(* Logix 5000 project; controller PLC_MCC1300_75F1 vendor 1 type 14 code 166 rev 32.11; software revision 32.04; part 4 of 83 *)
(* tags used below, declared in another part *)
   GP_AccTimeForGap : GP_AccTimeForGap;
   GP_CheckIdPlatePresent : GP_CheckIdPlatePresent;
   GP_ConversionXY : GP_ConversionXY;
   GP_ConvertDataFromStacker : GP_ConvertDataFromStacker;
   GP_ConvertDataToStacker : GP_ConvertDataToStacker;
   GP_InvertCapxLite : GP_InvertCapxLite;

ADD_ON_INSTRUCTION GP_AccTimeForGap   (* revision 1.0 *)
VAR_INPUT
   IN_dLehrSpeed_mm_min : DINT; {access None, required}
   IN_dLineSpeed_mm_min : DINT; {access None, required}
   IN_rAcc_m_s2 : REAL; {access None, required}
   IN_dGapRequested_cmm : DINT; {access None, required}
END_VAR
VAR_OUTPUT
   OUT_dAccTime_ms : DINT; {access None, required}
END_VAR
VAR
   TMP_rSpeed_mm_s : REAL; {access None}
   TMP_rConvSpeed_mm_s : REAL; {access None}
   TMP_rAccConv_mm_s2 : REAL; {access None}
   TMP_rAcc : REAL; {access None}
   TMP_rSv : REAL; {access None}
   TMP_dGap_mm : DINT; {access None}
END_VAR

ROUTINE Logic   (* structured text *)
   
   TMP_rSpeed_mm_s := (IN_dLehrSpeed_mm_min / 60.0);
   TMP_rConvSpeed_mm_s := (IN_dLineSpeed_mm_min / 60.0);
   TMP_rAccConv_mm_s2 := (IN_rAcc_m_s2 * 1000.0);
   TMP_dGap_mm := (IN_dGapRequested_cmm / 100);
   
   TMP_rAcc := ((TMP_rSpeed_mm_s*-1) + SQRT(TMP_rSpeed_mm_s**2 + (2*TMP_rAccConv_mm_s2*200)))/TMP_rAccConv_mm_s2;
   IF ((TMP_rAcc*TMP_rAccConv_mm_s2) + TMP_rSpeed_mm_s) > TMP_rConvSpeed_mm_s THEN
       TMP_rAcc := (TMP_rConvSpeed_mm_s - TMP_rSpeed_mm_s) / TMP_rAccConv_mm_s2;
       TMP_rSv := TMP_dGap_mm - (0.5*(TMP_rAcc**2)*TMP_rAccConv_mm_s2) - (TMP_rSpeed_mm_s*TMP_rAcc);
       TMP_rAcc := TMP_rAcc + (TMP_rSv/TMP_rConvSpeed_mm_s);
   END_IF;
   
   IF IN_dGapRequested_cmm > 0 THEN
       OUT_dAccTime_ms := TMP_rAcc * 1000.0;
   ELSE
       OUT_dAccTime_ms := 0;
   END_IF;
   
END_ROUTINE
END_ADD_ON_INSTRUCTION

ADD_ON_INSTRUCTION GP_BaricenterDefinition   (* revision 1.0 *)
VAR_INPUT
   In_dHeadPosition : DINT; {required}   // Head position on conveyor below [mm/100]
END_VAR
VAR_IN_OUT
   InOut_ConvoyData : UDT_Convoy_SL; {required}
END_VAR
VAR_INPUT
   In_dInLitePos : DINT; {access None, required}   // Position input lite - Left to Right line flow(0=AX; 1=XA)
   In_dOutDirection : DINT; {required}   // Direction of lateral flow (0=Left; 1=Right; 2=CW(rotation); 3=CCW(rotation))
   In_dOutLitePos : DINT; {access None, required}   // Position output lite - Left to Right line flow(0=AX; 1=XA)
   In_dOffset1 : DINT; {required}   // Distance of start conveyorIn and axe conveyorOut [mm/100]
   In_dOffset2 : DINT; {required}   // (NU)
   In_dConveyorLenght : DINT; {access None, required}   // Conveyor below [mm/100]
   In_dConveyorWidth : DINT; {access None, required}   // Conveyor below [mm/100]
END_VAR
VAR
   TMP_idxCap : DINT; {access None}
   TMP_IdxLite : DINT; {access None}
   TMP_MaxCap : DINT; {access None}
   TMP_MaxLite : DINT; {access None}
   TMP_d : DINT; {access None}
   TMP_NewBarycenterCap : DINT[10]; {access None}
   TMP_HeadPosition : DINT[10]; {access None}   // Head position cap [mm/100]
END_VAR

ROUTINE Logic   (* structured text *)
   ////////////////////////////////////////////////////////////
   //   Copyright (c)  <Key Automation srl>
   //------------------------------------------------------------
   //   Routine: GP_BaricenterDefinition - Logic
   //   Author: Gerto\admin
   //   Created: 2020-02-06
   //------------------------------------------------------------
   //   Description:
   //
   //
   //   History:
   //
   ////////////////////////////////////////////////////////////
   
   //Dimension array
   Size(InOut_ConvoyData.rgtCap,0,TMP_MaxCap);
   size(InOut_ConvoyData.rgtCap[0].rgtLite,0,TMP_MaxLite);
   
   //Conveyor deviation *****************************************
   
   //Cap1 Barycenter = HeadPosIn - 1/2 cap1lenght - offset1(distance between start of conveyorIn and exe of conveyorOut)
   //Cap2 Barycenter = Cap1 Barycenter - 1/2 Cap1Lenght - Gap - 1/2 Cap2Lenght
   //Cap3...
   if 	(In_dOutDirection = 0 and In_dInLitePos = 0 and In_dOutLitePos = 0) or
   	(In_dOutDirection = 0 and In_dInLitePos = 1 and In_dOutLitePos = 0) or
   	(In_dOutDirection = 1 and In_dInLitePos = 0 and In_dOutLitePos = 1) or
   	(In_dOutDirection = 1 and In_dInLitePos = 1 and In_dOutLitePos = 1) then
   	//Barycenter 1° cap
   	TMP_NewBarycenterCap[0] := In_dHeadPosition - InOut_ConvoyData.rgtCap[0].dLength_cmm/2 - In_dOffset1;
   	//Baricenter other caps
   	for TMP_idxCap := 1 to InOut_ConvoyData.dTotalCaps - 1 by 1 do
   		TMP_NewBarycenterCap[TMP_idxCap] := TMP_NewBarycenterCap[TMP_idxCap-1] - InOut_ConvoyData.rgtCap[TMP_idxCap-1].dLength_cmm / 2 - InOut_ConvoyData.rgtCap[TMP_idxCap-1].dReqGapForConv_cmm - InOut_ConvoyData.rgtCap[TMP_idxCap].dLength_cmm / 2;
   	end_for;
   end_if;
   
   
   //Cap1 Barycenter = - (head pos In - 1/2 Cap1Lenght - Offset1)
   //Cap2 Barycenter = Cap1 Barycenter + 1/2 Cap1Lenght + Gap + 1/2 Cap2Lenght-
   //Cap3...
   if 	(In_dOutDirection = 0 and In_dInLitePos = 0 and In_dOutLitePos = 1) or
   	(In_dOutDirection = 0 and In_dInLitePos = 1 and In_dOutLitePos = 1) or
   	(In_dOutDirection = 1 and In_dInLitePos = 0 and In_dOutLitePos = 0) or
   	(In_dOutDirection = 1 and In_dInLitePos = 1 and In_dOutLitePos = 0) then
   	//Baricenter 1° cap
   	TMP_NewBarycenterCap[0] := - (In_dHeadPosition - InOut_ConvoyData.rgtCap[0].dLength_cmm / 2 - In_dOffset1);
   	//Barycenter other caps
   	for TMP_idxCap := 1 to InOut_ConvoyData.dTotalCaps - 1 by 1 do
   		TMP_NewBarycenterCap[TMP_idxCap] := TMP_NewBarycenterCap[TMP_idxCap-1] + InOut_ConvoyData.rgtCap[TMP_idxCap-1].dLength_cmm / 2 + InOut_ConvoyData.rgtCap[TMP_idxCap-1].dReqGapForConv_cmm + InOut_ConvoyData.rgtCap[TMP_idxCap].dLength_cmm / 2;
   	end_for;
   end_if;
   
   
   //Rotator ****************************************************
   
   //Definition head position for all caps
   TMP_HeadPosition[0] := In_dHeadPosition;
   for TMP_idxCap := 1 to InOut_ConvoyData.dTotalCaps - 1 by 1 do
   	TMP_HeadPosition[TMP_idxCap] := TMP_HeadPosition[TMP_idxCap-1] - InOut_ConvoyData.rgtCap[TMP_idxCap-1].dLength_cmm - InOut_ConvoyData.rgtCap[TMP_idxCap-1].dReqGapForConv_cmm;
   end_for;
   
   
   //Cap[cap] Barycenter = (HeadPosCap[cap] - ConveyorLengthIn/2 - CapLength[cap]/2)
   if 	(In_dOutDirection = 2 and In_dInLitePos = 0 and In_dOutLitePos = 0) or
   	(In_dOutDirection = 3 and In_dInLitePos = 1 and In_dOutLitePos = 1) then
   	for TMP_idxCap := 0 to InOut_ConvoyData.dTotalCaps - 1 by 1 do
   		TMP_NewBarycenterCap[TMP_idxCap] := (TMP_HeadPosition[TMP_idxCap] - In_dConveyorLenght/2 - InOut_ConvoyData.rgtCap[TMP_idxCap].dLength_cmm/2);
   	end_for;
   end_if;
   
   //Cap[cap] Barycenter = - (HeadPosCap[cap] - ConveyorLengthIn/2 - CapLength[cap]/2)
   if 	(In_dOutDirection = 2 and In_dInLitePos = 1 and In_dOutLitePos = 1) or
   	(In_dOutDirection = 3 and In_dInLitePos = 0 and In_dOutLitePos = 0) then
   	for TMP_idxCap := 0 to InOut_ConvoyData.dTotalCaps - 1 by 1 do
   		TMP_NewBarycenterCap[TMP_idxCap] := -(TMP_HeadPosition[TMP_idxCap] - In_dConveyorLenght/2 - InOut_ConvoyData.rgtCap[TMP_idxCap].dLength_cmm/2);
   	end_for;
   end_if;
   
   //Write output
   for TMP_idxCap := 0 to InOut_ConvoyData.dTotalCaps - 1 by 1 do
   	for TMP_IdxLite := 0 to TMP_MaxLite - 1 by 1 do
   		if InOut_ConvoyData.rgtCap[TMP_idxCap].rgtLite[TMP_IdxLite].dID <> 0 then
   			InOut_ConvoyData.rgtCap[TMP_idxCap].rgtLite[TMP_IdxLite].dBarycenter_cmm := TMP_NewBarycenterCap[TMP_idxCap];
   		end_if;
   	end_for;
   end_for;
END_ROUTINE
END_ADD_ON_INSTRUCTION

ADD_ON_INSTRUCTION GP_CalculatePlateNumber   (* revision 1.0 *)
VAR_IN_OUT
   INO_tPlate : UDT_ConvoyCap_ZC; {required}   // Plate data
END_VAR
VAR
   TMP_dLiteSize : DINT; {access None}
   TMP_dLite : DINT; {access None}
   TMP_dCapSize : DINT; {access None}
   TMP_dCap : DINT; {access None}
   TMP_dCountCaps : DINT; {access None}
   TMP_dCountLites : DINT; {access None}
END_VAR

ROUTINE Logic   (* structured text *)
   //Initialize
   size(INO_tPlate.rgtCap[0],0,TMP_dCapSize);
   size(INO_tPlate.rgtCap[0].rgtLite[0],0,TMP_dLiteSize);
   
   TMP_dCountCaps:= 0;
   
   FOR TMP_dCap:= 0 TO TMP_dCapSize - 1 DO
   	TMP_dCountLites:= 0;
   	FOR TMP_dLite := 0 TO TMP_dLiteSize - 1 DO
   
   		IF INO_tPlate.rgtCap[TMP_dCap].rgtLite[TMP_dLite].dID <> 0 THEN
   
   			TMP_dCountLites := TMP_dCountLites +1 ;
   
   		END_IF;
   
   	END_FOR;
   
   	INO_tPlate.rgtCap[TMP_dCap].dNumLites := TMP_dCountLites ;
   
   	IF TMP_dCountLites > 0 THEN
   
   		TMP_dCountCaps := TMP_dCountCaps + 1 ;
   
   	END_IF;
   
   END_FOR;
   
   IF TMP_dCountCaps > 1 THEN
   
   	INO_tPlate.dTotalCaps := TMP_dCountCaps ;
   
   ELSE
   
   	INO_tPlate.dTotalCaps := 0 ;
   
   END_IF;
   
   EnableOut := 1 ;
END_ROUTINE
END_ADD_ON_INSTRUCTION

ADD_ON_INSTRUCTION GP_CheckIdAndDestination   (* revision 1.0 *)
VAR_INPUT
   IN_dDestMask1 : DINT; {access None, required}   // Destinations available on operator side
   IN_dDestMask2 : DINT; {access None, required}   // Destinations available on opposite operator side
END_VAR
VAR_IN_OUT
   INO_tPlate : UDT_Convoy_SL; {required}   // Plate data
   INO_rgxId : DINT[4]; {required}   // Array Id Plate present [Cap, Lite]
END_VAR
VAR_OUTPUT
   OUT_xIDPresent : BOOL; {access None}   // Id present
   OUT_xDest1Found : BOOL; {access None}   // Destinations found
   OUT_xDest2Found : BOOL; {access None}   // Destinations found
   OUT_xAlternative1Found : BOOL; {access None}   // Alternatives found
   OUT_xAlternative2Found : BOOL; {access None}   // Alternatives found
   OUT_x2Choice1Found : BOOL; {access None}   // 2°Choice found
   OUT_x2Choice2Found : BOOL; {access None}   // 2°Choice found
END_VAR
VAR
   TMP_dCap : DINT; {access None}
   TMP_dLite : DINT; {access None}
   TMP_dLiteSize : DINT; {access None}
   TMP_dCapSize : DINT; {access None}
END_VAR

ROUTINE Logic   (* structured text *)
   //Initialize
   INO_rgxId[0]:= 0; INO_rgxId[1]:= 0; INO_rgxId[2]:= 0;INO_rgxId[3]:= 0;
   OUT_xIDPresent:= 0;
   OUT_xDest1Found:= 0;
   OUT_xDest2Found:= 0;
   OUT_xAlternative1Found:= 0;
   OUT_xAlternative2Found:= 0;
   OUT_x2Choice1Found:= 0;
   OUT_x2Choice2Found:= 0;
   
   size(INO_tPlate.rgtCap[0],0,TMP_dCapSize);
   size(INO_tPlate.rgtCap[0].rgtLite[0],0,TMP_dLiteSize);
   
   //This function check ID Plate present
   //Max Cap = 4
   //Max Lite = 8
   FOR TMP_dCap:= 0 TO TMP_dCapSize - 1 DO
   
   	FOR TMP_dLite := 0 TO TMP_dLiteSize - 1 DO
   
   	IF INO_tPlate.rgtCap[TMP_dCap].rgtLite[TMP_dLite].dID <> 0 THEN
   
   		OUT_xIDPresent:= 1;
   		INO_rgxId[TMP_dCap].[TMP_dLite]:= 1;
   		//Find available destination
   		IF (INO_tPlate.rgtCap[TMP_dCap].rgtLite[TMP_dLite].tDestination.rgxMain AND IN_dDestMask1) > 0 THEN
   			OUT_xDest1Found:= 1;
   		ELSIF (INO_tPlate.rgtCap[TMP_dCap].rgtLite[TMP_dLite].tDestination.rgxMain AND IN_dDestMask2) > 0 THEN
   			OUT_xDest2Found:= 1;
   		ELSIF (INO_tPlate.rgtCap[TMP_dCap].rgtLite[TMP_dLite].tDestination.rgxAlternative AND IN_dDestMask1) > 0 THEN
   			OUT_xAlternative1Found:= 1;
   		ELSIF (INO_tPlate.rgtCap[TMP_dCap].rgtLite[TMP_dLite].tDestination.rgxAlternative AND IN_dDestMask2) > 0 THEN
   			OUT_xAlternative2Found:= 1;
   		ELSIF (INO_tPlate.rgtCap[TMP_dCap].rgtLite[TMP_dLite].tDestination.rgxSecChoice AND IN_dDestMask1) > 0 THEN
   			OUT_x2Choice1Found:= 1;
   		ELSIF (INO_tPlate.rgtCap[TMP_dCap].rgtLite[TMP_dLite].tDestination.rgxSecChoice AND IN_dDestMask2) > 0 THEN
   			OUT_x2Choice1Found:= 1;
   		END_IF;
   
   	END_IF;
   
   	END_FOR;
   
   END_FOR;
   
   EnableOut := 1 ;
END_ROUTINE
END_ADD_ON_INSTRUCTION

ADD_ON_INSTRUCTION GP_CheckIdPlatePresent   (* revision 1.0 *)
VAR_IN_OUT
   INO_tPlate : UDT_Convoy_SL; {required}   // Plate data
   INO_rgxId : DINT[10]; {required}   // Array Id Plate present [Cap, Lite]
END_VAR
VAR_OUTPUT
   OUT_xIDPresent : BOOL; {access None, required}   // Id present
   OUT_xDestToCheckPresent : BOOL; {access Read Only, required}
END_VAR
VAR_INPUT
   IN_DestToCheckPresence : DINT; {required}
END_VAR
VAR_OUTPUT
   OUT_dQtaLitesPresent : DINT;
END_VAR
VAR
   TMP_iCap : INT; {access None}
   TMP_iLite : INT; {access None}
   TMP_iLiteSize : INT; {access None}
   TMP_iCapSize : INT; {access None}
END_VAR

ROUTINE Logic   (* structured text *)
   //Initialize
   TMP_iCap:= 0; TMP_iLite:= 0;
   OUT_xIDPresent:= 0;
   OUT_xDestToCheckPresent := 0;
   INO_rgxId[0]:= 0; INO_rgxId[1]:= 0; INO_rgxId[2]:= 0;INO_rgxId[3]:= 0;
   OUT_dQtaLitesPresent := 0;
   
   size(INO_tPlate.rgtCap[0],0,TMP_iCapSize);
   size(INO_tPlate.rgtCap[0].rgtLite[0],0,TMP_iLiteSize);
   
   //This function check ID Plate present
   FOR TMP_iCap:= 0 TO TMP_iCapSize - 1 DO
   
   	FOR TMP_iLite := 0 TO TMP_iLiteSize - 1 DO
   
   	IF INO_tPlate.rgtCap[TMP_iCap].rgtLite[TMP_iLite].dID <> 0 THEN
   		OUT_dQtaLitesPresent := OUT_dQtaLitesPresent +1;
   		OUT_xIDPresent:= 1;
   		INO_rgxId[TMP_iCap].[TMP_iLite]:= 1;
   		if  INO_tPlate.rgtCap[TMP_iCap].rgtLite[TMP_iLite].tDestination.rgxMain.[IN_DestToCheckPresence] then
   			OUT_xDestToCheckPresent := 1;
   		end_if;
   
   	END_IF;
   
   	END_FOR;
   
   END_FOR;
   
   EnableOut := 1 ;
END_ROUTINE
END_ADD_ON_INSTRUCTION

ADD_ON_INSTRUCTION GP_CheckSnapIndex   (* revision 1.0 *)
VAR_IN_OUT
   INO_rgtTrackingSearch : GP_TrackingSearchPlate_STC; {required}
   INO_rgtBufferPlate : UDT_LINE_BUFFER_PLATE; {required}
END_VAR
VAR_OUTPUT
   OUT_dIndex : DINT; {access None, required}
END_VAR
VAR
   TMP_dIndex : DINT; {access None}
   TMP_dPointer : DINT; {access None}
END_VAR

ROUTINE Logic   (* structured text *)
   
   OUT_dIndex := 0;
   FOR TMP_dIndex := 0 TO 4 DO
   	TMP_dPointer := INO_rgtTrackingSearch.rgdHeadPointer[TMP_dIndex];
   	IF TMP_dPointer > 0 THEN
   		IF INO_rgtBufferPlate.rgtPlate[TMP_dPointer].tData.rgtCap[0].dNumLites > 1 THEN
   			OUT_dIndex := INO_rgtTrackingSearch.rgdHeadPointer[TMP_dIndex];
   			EXIT;
   		END_IF;
   	END_IF;
   END_FOR;
   
END_ROUTINE
END_ADD_ON_INSTRUCTION

ADD_ON_INSTRUCTION GP_CompactConvoy   (* revision 1.0 *)
VAR_IN_OUT
   InOut_ConvoyData : UDT_Convoy_SL; {required}
   Const_ConvoyData_Empty : UDT_Convoy_SL; {constant, required}
END_VAR
VAR
   TMP_MaxCap : DINT; {access None}
   TMP_MaxLite : DINT; {access None}
   TMP_d : DINT; {access None}
   TMP_idxCap : DINT; {access None}
   TMP_idxLite : DINT; {access None}
   TMP_FirstCapFinded : DINT; {access None}
   TMP_LastCapFinded : DINT; {access None}
END_VAR

ROUTINE Logic   (* structured text *)
   ////////////////////////////////////////////////////////////
   //   Copyright (c)  <Key Automation srl>
   //------------------------------------------------------------
   //   Routine: GP_CompactConvoy - Logic
   //   Author: Gerto\admin
   //   Created: 2020-02-03
   //------------------------------------------------------------
   //   Description:
   //
   //
   //   History:
   //
   ////////////////////////////////////////////////////////////
   
   //Dimension array
   Size(InOut_ConvoyData.rgtCap,0,TMP_MaxCap);
   size(InOut_ConvoyData.rgtCap[0].rgtLite,0,TMP_MaxLite);
   
   //Init
   TMP_FirstCapFinded := -1;
   TMP_LastCapFinded := 99;
   
   
   //Find first cap present before compacting
   for TMP_idxCap := 0 to TMP_MaxCap-1 by 1 do
   	for TMP_idxLite := 0 to TMP_MaxLite-1 by 1 do
   		if InOut_ConvoyData.rgtCap[TMP_idxCap].rgtLite[TMP_idxLite].dID <> 0 then
   			TMP_FirstCapFinded := TMP_idxCap;
   			exit;
   		end_if;
   	end_for;
   	if TMP_FirstCapFinded >= 0 then
   		exit;
   	end_if;
   end_for;
   
   
   //Move first cap present to start array and so on...
   If TMP_FirstCapFinded > 0 then
   	for TMP_idxCap := 0 to TMP_MaxCap-1 by 1 do
   		if TMP_FirstCapFinded+TMP_idxCap <= TMP_MaxCap-1 then
   			cop(InOut_ConvoyData.rgtCap[TMP_FirstCapFinded+TMP_idxCap],InOut_ConvoyData.rgtCap[TMP_idxCap],1);
   			cop(Const_ConvoyData_Empty.rgtCap[0],InOut_ConvoyData.rgtCap[TMP_FirstCapFinded+TMP_idxCap],1);
   		end_if;
   	end_for;
   end_if;
   
   //Find last cap(with lite ID) on convoy after compacting
   for TMP_idxCap := TMP_MaxCap-1 to 0 by -1 do
   	for TMP_idxLite := 0 to TMP_MaxLite-1 by +1 do
   		if InOut_ConvoyData.rgtCap[TMP_idxCap].rgtLite[TMP_idxLite].dID <> 0 then
   			TMP_LastCapFinded := TMP_idxCap;
   			exit;
   		end_if;
   	end_for;
   	if TMP_LastCapFinded <= TMP_MaxCap-1 then
   		exit;
   	end_if;
   end_for;
   
   //Clear data cap starting from last cap present till the end of array
   if TMP_LastCapFinded < TMP_MaxCap-1 then
   	for TMP_idxCap := TMP_LastCapFinded+1 to TMP_MaxCap-1 by 1 do
   		cop(Const_ConvoyData_Empty.rgtCap[0],InOut_ConvoyData.rgtCap[TMP_idxCap],1);
   	end_for;
   end_if;
   
   
   //Write General convoy data
   
   //Convoy length
   TMP_d := 0;
   if TMP_LastCapFinded <= TMP_MaxCap-1 then
   	for TMP_idxCap := 0 to TMP_LastCapFinded by 1 do
   		TMP_d:= TMP_d + InOut_ConvoyData.rgtCap[TMP_idxCap].dLength_cmm;
   	end_for;
   end_if;
   TMP_d := TMP_d + TMP_LastCapFinded * InOut_ConvoyData.dGapCaps_cmm;
   InOut_ConvoyData.dLength_cmm := TMP_d;
   
   //Qta Cap
   InOut_ConvoyData.dTotalCaps := TMP_LastCapFinded + 1;
END_ROUTINE
END_ADD_ON_INSTRUCTION

ADD_ON_INSTRUCTION GP_CompactConvoy_V2   (* revision 1.0 *)
VAR_IN_OUT
   InOut_ConvoyData : UDT_Convoy_SL; {required}
   Const_ConvoyData_Empty : UDT_Convoy_SL; {constant, required}
END_VAR
VAR
   TMP_MaxCap : DINT; {access None}
   TMP_MaxLite : DINT; {access None}
   TMP_d : DINT; {access None}
   TMP_idxCap : DINT; {access None}
   TMP_idxLite : DINT; {access None}
   TMP_CapPresent : BOOL; {access None}
   TMP_CapPrecPresent : BOOL; {access None}
END_VAR

ROUTINE Logic   (* structured text *)
   ////////////////////////////////////////////////////////////
   //   Copyright (c)  <Key Automation srl>
   //------------------------------------------------------------
   //   Routine: GP_CompactConvoy - Logic
   //   Author: Gerto\admin
   //   Created: 2020-02-03
   //------------------------------------------------------------
   //   Description:
   //
   //
   //   History:
   //
   ////////////////////////////////////////////////////////////
   
   //Dimension array
   Size(InOut_ConvoyData.rgtCap,0,TMP_MaxCap);
   size(InOut_ConvoyData.rgtCap[0].rgtLite,0,TMP_MaxLite);
   
   //Compact caps to start array
   for TMP_idxCap := 1 to TMP_MaxCap - 1 by 1 do
   	TMP_CapPrecPresent := 0;
   	TMP_CapPresent := 0;
   	for TMP_idxLite := 0 to TMP_MaxLite -1 by 1 do
   		if InOut_ConvoyData.rgtCap[TMP_idxCap-1].rgtLite[TMP_idxLite].dID <> 0 then
   			TMP_CapPrecPresent := 1;
   			exit;
   		end_if;
   	end_for;
   	for TMP_idxLite := 0 to TMP_MaxLite -1 by 1 do
   		if InOut_ConvoyData.rgtCap[TMP_idxCap].rgtLite[TMP_idxLite].dID <> 0 then
   			TMP_CapPresent := 1;
   			exit;
   		end_if;
   	end_for;
   	if not TMP_CapPrecPresent and TMP_CapPresent then
   		cop(InOut_ConvoyData.rgtCap[TMP_idxCap],InOut_ConvoyData.rgtCap[TMP_idxCap-1],1);
   		cop(Const_ConvoyData_Empty.rgtCap[0],InOut_ConvoyData.rgtCap[TMP_idxCap],1);
   		TMP_idxCap := TMP_idxCap -1;
   	end_if;
   end_for;
   
   //Qta Caps
   InOut_ConvoyData.dTotalCaps := 0;
   for TMP_idxCap := 0 to TMP_MaxCap - 1 by 1 do
   	for TMP_idxLite := 0 to TMP_MaxLite -1 by 1 do
   		if InOut_ConvoyData.rgtCap[TMP_idxCap].rgtLite[TMP_idxLite].dID <> 0 then
   			InOut_ConvoyData.dTotalCaps := InOut_ConvoyData.dTotalCaps + 1;
   			exit;
   		end_if;
   	end_for;
   end_for;
   
   //Convoy length
   for TMP_idxCap := 0 to InOut_ConvoyData.dTotalCaps - 1 by 1 do
   	InOut_ConvoyData.dLength_cmm := InOut_ConvoyData.dLength_cmm + InOut_ConvoyData.rgtCap[TMP_idxCap].dLength_cmm;
   	if TMP_idxCap < InOut_ConvoyData.dTotalCaps - 1 then
   		InOut_ConvoyData.dLength_cmm := InOut_ConvoyData.dLength_cmm + InOut_ConvoyData.rgtCap[TMP_idxCap].dReqGapForConv_cmm;
   	end_if;
   end_for;
   
END_ROUTINE
END_ADD_ON_INSTRUCTION

ADD_ON_INSTRUCTION GP_ConversionXY   (* revision 1.0 *)
VAR_INPUT
   IN_rXvalue : REAL; {access None, required}   // Input value X
   IN_rXmin : REAL; {access None, required}   // Minimum value X
   IN_rXmax : REAL; {access None, required}   // Maximum value X
   IN_rYmin : REAL; {access None, required}   // Minimum value Y
   IN_rYmax : REAL; {access None, required}   // Maximum value Y
END_VAR
VAR_OUTPUT
   OUT_rYvalue : REAL; {access None, required}   // Output value Y
END_VAR
VAR
   TMP_rDelta_y : REAL; {access None}
   TMP_rDelta_x : REAL; {access None}
END_VAR

ROUTINE Logic   (* structured text *)
   
   //Inizialize Output
   OUT_rYvalue := 0.0;
   
   //    (S_x -Xmin)*(Ymax-Ymin)
   //S_y=------------------------ + Ymin
   //         (Xmax-Xmin)
   
   TMP_rDelta_x := IN_rXmax - IN_rXmin;
   TMP_rDelta_y := IN_rYmax - IN_rYmin;
   
   IF IN_rXmax <> IN_rXmin THEN
     OUT_rYvalue := (((IN_rXvalue - IN_rXmin) * TMP_rDelta_y) / TMP_rDelta_x) + IN_rYmin;
   ELSE
     OUT_rYvalue := 0.0;
   END_IF;
   
END_ROUTINE
END_ADD_ON_INSTRUCTION

ADD_ON_INSTRUCTION GP_ConvertDataFromStacker   (* revision 1.0 *)
VAR_IN_OUT
   In_tStkData : UDT_PlateData_Convoy; {required}
   Out_tConvoyData : UDT_Convoy_SL; {required}
END_VAR
VAR_INPUT
   In_GapBetweenLites : DINT; {access None}
END_VAR
VAR
   TMP_LiteAPresent : BOOL; {access None}
   TMP_LiteBPresent : BOOL; {access None}
   TMP_Idx_Lite : DINT; {access None}
   TMP_Idx_Pos : DINT; {access None}   // [0=Right; 1=Left]
   TMP_x : BOOL; {access None}
END_VAR

ROUTINE Logic   (* structured text *)
   ////////////////////////////////////////////////////////////
   //   Copyright (c)  <Key Automation srl>
   //------------------------------------------------------------
   //   Routine: GP_ConvertDataToStacker - Logic
   //   Author: Gerto\admin
   //   Created: 2020-02-10
   //------------------------------------------------------------
   //   Description:
   //
   //
   //   History:
   //
   ////////////////////////////////////////////////////////////
   
   //Set presence lites
   TMP_LiteAPresent := In_tStkData.tLite[0].dID <> 0;
   TMP_LiteBPresent := In_tStkData.tLite[1].dID <> 0;
   
   //Convoy data
   Out_tConvoyData.dLength_cmm := In_tStkData.dTotLenght_cmm;
   Out_tConvoyData.rgtCap[0].dWidth_cmm := In_tStkData.dTotWidth_cmm;
   
   //Lite Data
   
   //Both lites
   If TMP_LiteAPresent and TMP_LiteBPresent then
   	For TMP_Idx_Lite := 0 to 1 by 1 do
   		TMP_Idx_Pos := TMP_Idx_Lite;
   		Out_tConvoyData.rgtCap[0].rgtLite[TMP_Idx_Lite].dID := In_tStkData.tLite[TMP_Idx_Pos].dID;
   		Out_tConvoyData.rgtCap[0].rgtLite[TMP_Idx_Lite].dProductionID := In_tStkData.tLite[TMP_Idx_Pos].dProduction_ID;
   		Out_tConvoyData.rgtCap[0].dLength_cmm := In_tStkData.tLite[TMP_Idx_Pos].dLenght_cmm;
   		Out_tConvoyData.rgtCap[0].rgtLite[TMP_Idx_Lite].dWidth_cmm := In_tStkData.tLite[TMP_Idx_Pos].dWidth_cmm;
   		Out_tConvoyData.rgtCap[0].dThickness_cmm := In_tStkData.tLite[TMP_Idx_Pos].dThick_cmm;
   		Out_tConvoyData.rgtCap[0].rgtLite[TMP_Idx_Lite].tDestination.rgxMain := In_tStkData.tLite[TMP_Idx_Pos].rgxMain;
   		Out_tConvoyData.rgtCap[0].rgtLite[TMP_Idx_Lite].tDestination.rgxAlternative := In_tStkData.tLite[TMP_Idx_Pos].rgxAlternative;
   		Out_tConvoyData.rgtCap[0].dID := In_tStkData.tLite[TMP_Idx_Pos].dID;
   		Out_tConvoyData.rgtCap[0].dNumLites := 2;
   		Out_tConvoyData.dTotalCaps := 1;
   		Out_tConvoyData.rgtCap[0].rgtLite[0].dBarycenter_cmm := - (Out_tConvoyData.rgtCap[0].rgtLite[TMP_Idx_Lite].dWidth_cmm / 2 + In_GapBetweenLites);
   		Out_tConvoyData.rgtCap[0].rgtLite[1].dBarycenter_cmm := Out_tConvoyData.rgtCap[0].rgtLite[TMP_Idx_Lite].dWidth_cmm / 2 + In_GapBetweenLites;
   	end_for;
   end_if;
   
   //Any single case
   TMP_x := 0;
   If TMP_LiteAPresent and not TMP_LiteBPresent then //and In_tStkData.dPositionLite = 1  then
   	TMP_Idx_Lite := 0;
   	TMP_Idx_Pos := 0;
   	TMP_x := 1;
   //elsif TMP_LiteAPresent and not TMP_LiteBPresent then //and In_tStkData.dPositionLite = 2 then//
   //	TMP_Idx_Lite := 0;
   //	TMP_Idx_Pos := 1;
   //	TMP_x := 1;
   //elsif not TMP_LiteAPresent and TMP_LiteBPresent then //and In_tStkData.dPositionLite = 1 then//
   //	TMP_Idx_Lite := 1;
   //	TMP_Idx_Pos := 0;
   //	TMP_x := 1;
   elsif not TMP_LiteAPresent and TMP_LiteBPresent then //and In_tStkData.dPositionLite = 2 then
   	TMP_Idx_Lite := 1;
   	TMP_Idx_Pos := 1;
   	TMP_x := 1;
   end_if;
   
   if TMP_x then
   	TMP_Idx_Pos := TMP_Idx_Lite;
   	Out_tConvoyData.rgtCap[0].rgtLite[TMP_Idx_Lite].dID := In_tStkData.tLite[TMP_Idx_Pos].dID;
   	Out_tConvoyData.rgtCap[0].rgtLite[TMP_Idx_Lite].dProductionID := In_tStkData.tLite[TMP_Idx_Pos].dProduction_ID;
   	Out_tConvoyData.rgtCap[0].dLength_cmm := In_tStkData.tLite[TMP_Idx_Pos].dLenght_cmm;
   	Out_tConvoyData.rgtCap[0].rgtLite[TMP_Idx_Lite].dWidth_cmm := In_tStkData.tLite[TMP_Idx_Pos].dWidth_cmm;
   	Out_tConvoyData.rgtCap[0].dThickness_cmm := In_tStkData.tLite[TMP_Idx_Pos].dThick_cmm;
   	Out_tConvoyData.rgtCap[0].rgtLite[TMP_Idx_Lite].tDestination.rgxMain := In_tStkData.tLite[TMP_Idx_Pos].rgxMain;
   	Out_tConvoyData.rgtCap[0].rgtLite[TMP_Idx_Lite].tDestination.rgxAlternative := In_tStkData.tLite[TMP_Idx_Pos].rgxAlternative;
   	Out_tConvoyData.rgtCap[0].dID := In_tStkData.tLite[TMP_Idx_Pos].dID;
   	Out_tConvoyData.rgtCap[0].dNumLites := 1;
   	Out_tConvoyData.dTotalCaps := 1;
   	if In_tStkData.dFormat = 1 then
   		Out_tConvoyData.rgtCap[0].rgtLite[0].dBarycenter_cmm := 0;
   	elsif TMP_Idx_Lite = 0 then
   		Out_tConvoyData.rgtCap[0].rgtLite[0].dBarycenter_cmm := - (Out_tConvoyData.rgtCap[0].rgtLite[TMP_Idx_Lite].dWidth_cmm / 2 + In_GapBetweenLites);
   	elsif	 TMP_Idx_Lite = 1 then
   		Out_tConvoyData.rgtCap[0].rgtLite[1].dBarycenter_cmm := Out_tConvoyData.rgtCap[0].rgtLite[TMP_Idx_Lite].dWidth_cmm / 2 + In_GapBetweenLites;
   	end_if;
   
   end_if;
END_ROUTINE
END_ADD_ON_INSTRUCTION

ADD_ON_INSTRUCTION GP_ConvertDataToStacker   (* revision 1.0 *)
VAR_IN_OUT
   In_tConvoyData : UDT_Convoy_SL; {required}
   Out_tStkData : UDT_PlateData_Convoy; {required}
END_VAR
VAR
   TMP_LiteAPresent : BOOL; {access None}
   TMP_LiteBPresent : BOOL; {access None}
   TMP_Idx_Lite : DINT; {access None}
   TMP_Idx_Pos : DINT; {access None}   // [0=Right; 1=Left]
   TMP_x : BOOL; {access None}
END_VAR

ROUTINE Logic   (* structured text *)
   ////////////////////////////////////////////////////////////
   //   Copyright (c)  <Key Automation srl>
   //------------------------------------------------------------
   //   Routine: GP_ConvertDataToStacker - Logic
   //   Author: Gerto\admin
   //   Created: 2020-02-10
   //------------------------------------------------------------
   //   Description:
   //
   //
   //   History:
   //
   ////////////////////////////////////////////////////////////
   
   
   //Init
   for TMP_Idx_Pos := 0 to 1 by 1 do
   	Out_tStkData.tLite[TMP_Idx_Pos].dID := 0;
   	Out_tStkData.tLite[TMP_Idx_Pos].dProduction_ID := 0;
   	Out_tStkData.tLite[TMP_Idx_Pos].dLenght_cmm := 0;
   	Out_tStkData.tLite[TMP_Idx_Pos].dWidth_cmm := 0;
   	Out_tStkData.tLite[TMP_Idx_Pos].dThick_cmm := 0;
   	Out_tStkData.tLite[TMP_Idx_Pos].rgxOrigin := 0;
   	Out_tStkData.tLite[TMP_Idx_Pos].rgxMain := 0;
   	Out_tStkData.tLite[TMP_Idx_Pos].rgxAlternative := 0;
   	Out_tStkData.tLite[TMP_Idx_Pos].xCoated := 0;
   	Out_tStkData.tLite[TMP_Idx_Pos].xCoverPlate := 0;
   end_for;
   
   //Set presence lites
   TMP_LiteAPresent := In_tConvoyData.rgtCap[0].rgtLite[0].dID <> 0;
   TMP_LiteBPresent := In_tConvoyData.rgtCap[0].rgtLite[1].dID <> 0;
   
   //Convoy data
   Out_tStkData.dIDTx := In_tConvoyData.rgtCap[0].rgtLite[0].dID;
   if Out_tStkData.dIDTx = 0 then
   	Out_tStkData.dIDTx := In_tConvoyData.rgtCap[0].rgtLite[1].dID;
   end_if;
   Out_tStkData.dTotLenght_cmm := In_tConvoyData.dLength_cmm;
   Out_tStkData.dTotWidth_cmm := In_tConvoyData.rgtCap[0].dWidth_cmm;
   
   //Out_tStkData.dFormat := 2;
   //if In_tConvoyData.rgtCap[0].rgtLite[0].dWidth_cmm > In_MaxLiteWidththen//
   //	Out_tStkData.dFormat := 1;
   //end_if;
   
   Out_tStkData.dNumLites := In_tConvoyData.rgtCap[0].dNumLites;
   
   
   Out_tStkData.dPositionLite := 0;
   Out_tStkData.dFormat := 1;
   if  (TMP_LiteAPresent and not TMP_LiteBPresent) or
   	(Not TMP_LiteAPresent and TMP_LiteBPresent) then
   		if  (TMP_LiteAPresent and In_tConvoyData.rgtCap[0].rgtLite[0].dBarycenter_cmm < 0) or
   			(TMP_LiteBPresent and In_tConvoyData.rgtCap[0].rgtLite[1].dBarycenter_cmm < 0) then
   				Out_tStkData.dPositionLite := 1;
   				Out_tStkData.dFormat := 2;
   		end_if;
   		if  (TMP_LiteAPresent and In_tConvoyData.rgtCap[0].rgtLite[0].dBarycenter_cmm > 0) or
   			(TMP_LiteBPresent and In_tConvoyData.rgtCap[0].rgtLite[1].dBarycenter_cmm > 0) then
   				Out_tStkData.dPositionLite := 2;
   				Out_tStkData.dFormat := 2;
   		end_if;
   elsif TMP_LiteAPresent and TMP_LiteBPresent then
   	Out_tStkData.dFormat := 2;
   end_if;
   
   //Lite Data
   
   //Both lites
   If TMP_LiteAPresent and TMP_LiteBPresent then
   	For TMP_Idx_Lite := 0 to 1 by 1 do
   		TMP_Idx_Pos := TMP_Idx_Lite;
   		Out_tStkData.tLite[TMP_Idx_Pos].dID := In_tConvoyData.rgtCap[0].rgtLite[TMP_Idx_Lite].dID;
   		Out_tStkData.tLite[TMP_Idx_Pos].dProduction_ID := In_tConvoyData.rgtCap[0].rgtLite[TMP_Idx_Lite].dProductionID;
   		Out_tStkData.tLite[TMP_Idx_Pos].dLenght_cmm := In_tConvoyData.rgtCap[0].dLength_cmm;
   		Out_tStkData.tLite[TMP_Idx_Pos].dWidth_cmm := In_tConvoyData.rgtCap[0].rgtLite[TMP_Idx_Lite].dWidth_cmm;
   		Out_tStkData.tLite[TMP_Idx_Pos].dThick_cmm := In_tConvoyData.rgtCap[0].dThickness_cmm;
   		Out_tStkData.tLite[TMP_Idx_Pos].rgxOrigin := 0;
   		Out_tStkData.tLite[TMP_Idx_Pos].rgxMain := In_tConvoyData.rgtCap[0].rgtLite[TMP_Idx_Lite].tDestination.rgxMain;
   		Out_tStkData.tLite[TMP_Idx_Pos].rgxAlternative := In_tConvoyData.rgtCap[0].rgtLite[TMP_Idx_Lite].tDestination.rgxAlternative;
   		Out_tStkData.tLite[TMP_Idx_Pos].xCoated := 0;
   		Out_tStkData.tLite[TMP_Idx_Pos].xCoverPlate := 0;
   	end_for;
   end_if;
   
   //Any single case
   TMP_x := 0;
   If TMP_LiteAPresent and not TMP_LiteBPresent and Out_tStkData.dPositionLite <= 1  then
   	TMP_Idx_Lite := 0;
   	TMP_Idx_Pos := 0;
   	TMP_x := 1;
   elsif TMP_LiteAPresent and not TMP_LiteBPresent and Out_tStkData.dPositionLite = 2 then
   	TMP_Idx_Lite := 0;
   	TMP_Idx_Pos := 1;
   	TMP_x := 1;
   elsif not TMP_LiteAPresent and TMP_LiteBPresent and Out_tStkData.dPositionLite <= 1 then
   	TMP_Idx_Lite := 1;
   	TMP_Idx_Pos := 0;
   	TMP_x := 1;
   elsif not TMP_LiteAPresent and TMP_LiteBPresent and Out_tStkData.dPositionLite = 2 then
   	TMP_Idx_Lite := 1;
   	TMP_Idx_Pos := 1;
   	TMP_x := 1;
   end_if;
   
   if TMP_x then
   	Out_tStkData.tLite[TMP_Idx_Pos].dID := In_tConvoyData.rgtCap[0].rgtLite[TMP_Idx_Lite].dID;
   	Out_tStkData.tLite[TMP_Idx_Pos].dProduction_ID := In_tConvoyData.rgtCap[0].rgtLite[TMP_Idx_Lite].dProductionID;
   	Out_tStkData.tLite[TMP_Idx_Pos].dLenght_cmm := In_tConvoyData.rgtCap[0].dLength_cmm;
   	Out_tStkData.tLite[TMP_Idx_Pos].dWidth_cmm := In_tConvoyData.rgtCap[0].rgtLite[TMP_Idx_Lite].dWidth_cmm;
   	Out_tStkData.tLite[TMP_Idx_Pos].dThick_cmm := In_tConvoyData.rgtCap[0].dThickness_cmm;
   	Out_tStkData.tLite[TMP_Idx_Pos].rgxOrigin := 0;
   	Out_tStkData.tLite[TMP_Idx_Pos].rgxMain := In_tConvoyData.rgtCap[0].rgtLite[TMP_Idx_Lite].tDestination.rgxMain;
   	Out_tStkData.tLite[TMP_Idx_Pos].rgxAlternative := In_tConvoyData.rgtCap[0].rgtLite[TMP_Idx_Lite].tDestination.rgxAlternative;
   	Out_tStkData.tLite[TMP_Idx_Pos].xCoated := 0;
   	Out_tStkData.tLite[TMP_Idx_Pos].xCoverPlate := 0;
   end_if;
END_ROUTINE
END_ADD_ON_INSTRUCTION

ADD_ON_INSTRUCTION GP_GetIdFromData   (* revision 1.0 *)
VAR_IN_OUT
   INO_tPlate : UDT_Convoy_SL; {required}   // Plate data
END_VAR
VAR_OUTPUT
   OUT_dID : DINT; {access None}   // Id Plate
   OUT_dIdProduction : DINT; {access None}   // Id Production
END_VAR
VAR
   TMP_dCap : DINT; {access None}
   TMP_dLite : DINT; {access None}
   TMP_dLiteSize : DINT; {access None}
   TMP_dCapSize : DINT; {access None}
END_VAR

ROUTINE Logic   (* structured text *)
   //Initialize
   TMP_dCap:= 0; TMP_dLite:= 0;
   OUT_dIdProduction:= 0;
   OUT_dID:= 0;
   
   size(INO_tPlate.rgtCap[0],0,TMP_dCapSize);
   size(INO_tPlate.rgtCap[0].rgtLite[0],0,TMP_dLiteSize);
   
   FOR TMP_dCap:= 0 TO TMP_dCapSize - 1 DO
   
   	FOR TMP_dLite := 0 TO TMP_dLiteSize - 1 DO
   
   	IF INO_tPlate.rgtCap[TMP_dCap].rgtLite[TMP_dLite].dID <> 0 AND INO_tPlate.rgtCap[TMP_dCap].rgtLite[TMP_dLite].dProductionID <> 0 THEN
   
   		OUT_dIdProduction:= INO_tPlate.rgtCap[TMP_dCap].rgtLite[TMP_dLite].dProductionID;
   		OUT_dID:= INO_tPlate.rgtCap[TMP_dCap].rgtLite[TMP_dLite].dID;
   		TND();
   
   	END_IF;
   
   	END_FOR;
   
   END_FOR;
   
   EnableOut := 1 ;
END_ROUTINE
END_ADD_ON_INSTRUCTION
